(* Logix 5000 project; controller MV vendor 1 type 14 code 217 rev 31.11; software revision 31.00; part 20 of 53 *)
(* tags used below, declared in another part *)
   CheckTimeMask : INT;
   CWD : CHECKWORD_FLAGS;
   Delphi_Does_Eng_Func : BOOL;
   MC_CH1_DR2 : PlantItem;   // CH1_DR2
   MC_CH1_DT1 : PlantItem;   // CH1_DT1
   MC_CH1_DT2 : PlantItem;   // CH1_DT2
   MC_CH1_LF1 : PlantItem;   // CH1_LF1
   MC_CH1_PR1 : PlantItem;   // CH1_PR1
   MC_CH2_R1 : PlantItem;   // CH2_R1
   MC_CH2_R1R : PlantItem;   // CH2_R1R
   MC_CH2_R2 : PlantItem;   // CH2_R2
   MC_CH2_R2R : PlantItem;   // CH2_R2R
   MC_CH2_R3 : PlantItem;   // CH2_R3
   MC_CH2_R4 : PlantItem;   // CH2_R4
   MC_CH2_R5 : PlantItem;   // CH2_R5
   MC_CH2_R6 : PlantItem;   // CH2_R6
   MC_N255 : INT[255];   // CHECKWORDS Plant item checkword s
   TempChecktime : DINT;
(* MC_Common, continued *)

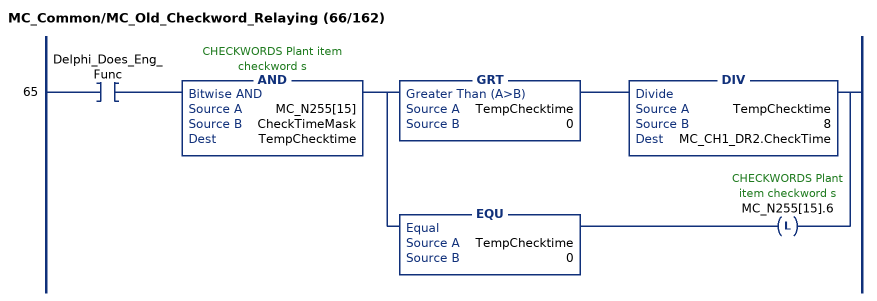
   [picture p337: MC_Common/MC_Old_Checkword_Relaying rungs 65-65]
   65: XIC(Delphi_Does_Eng_Func)AND(MC_N255[15],CheckTimeMask,TempChecktime)[GRT(TempChecktime,0) DIV(TempChecktime,8,MC_CH1_DR2.CheckTime) ,EQU(TempChecktime,0) OTL(MC_N255[15].6) ];
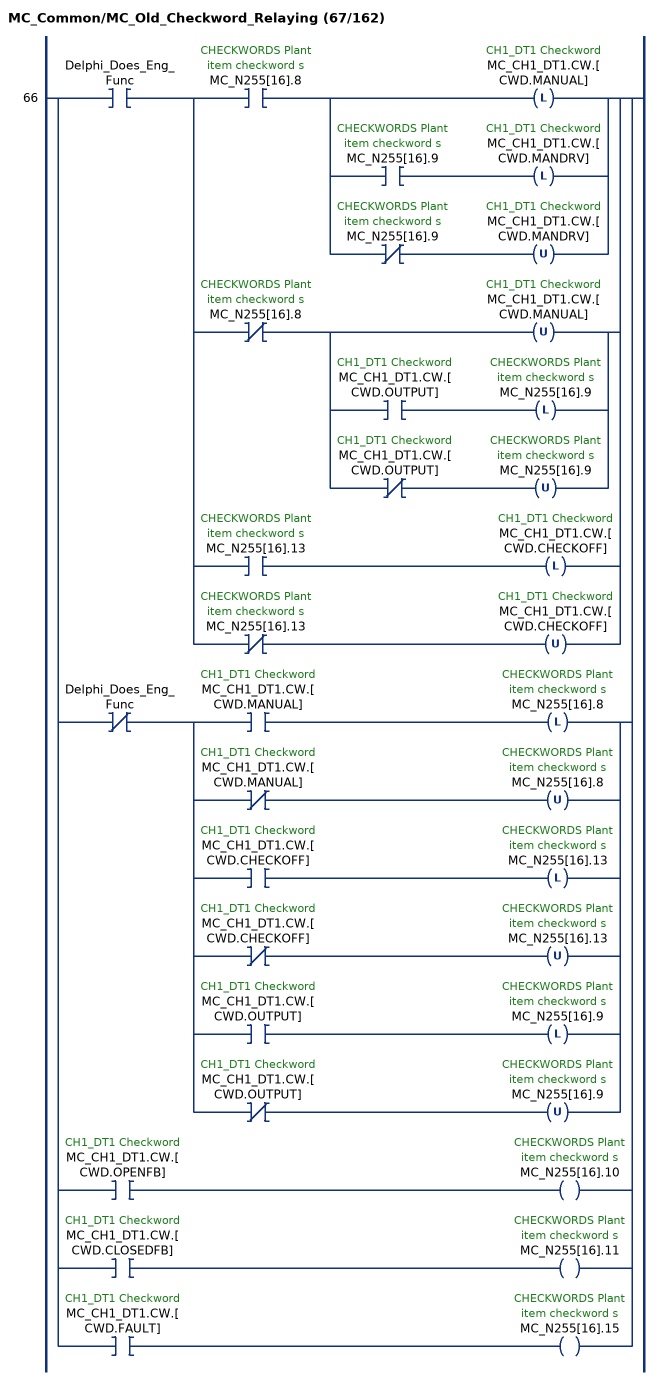
   66: [XIC(Delphi_Does_Eng_Func) [[XIC(MC_N255[16].8) [OTL(MC_CH1_DT1.CW.[CWD.MANUAL]) ,XIC(MC_N255[16].9) OTL(MC_CH1_DT1.CW.[CWD.MANDRV]) ,XIO(MC_N255[16].9) OTU(MC_CH1_DT1.CW.[CWD.MANDRV]) ] ,XIO(MC_N255[16].8) [OTU(MC_CH1_DT1.CW.[CWD.MANUAL]) ,[XIC(MC_CH1_DT1.CW.[CWD.OUTPUT]) OTL(MC_N255[16].9) ,XIO(MC_CH1_DT1.CW.[CWD.OUTPUT]) OTU(MC_N255[16].9) ] ] ] ,[XIC(MC_N255[16].13) OTL(MC_CH1_DT1.CW.[CWD.CHECKOFF]) ,XIO(MC_N255[16].13) OTU(MC_CH1_DT1.CW.[CWD.CHECKOFF]) ] ] ,XIO(Delphi_Does_Eng_Func) [[XIC(MC_CH1_DT1.CW.[CWD.MANUAL]) OTL(MC_N255[16].8) ,XIO(MC_CH1_DT1.CW.[CWD.MANUAL]) OTU(MC_N255[16].8) ] ,[XIC(MC_CH1_DT1.CW.[CWD.CHECKOFF]) OTL(MC_N255[16].13) ,XIO(MC_CH1_DT1.CW.[CWD.CHECKOFF]) OTU(MC_N255[16].13) ] ,[XIC(MC_CH1_DT1.CW.[CWD.OUTPUT]) OTL(MC_N255[16].9) ,XIO(MC_CH1_DT1.CW.[CWD.OUTPUT]) OTU(MC_N255[16].9) ] ] ,XIC(MC_CH1_DT1.CW.[CWD.OPENFB]) OTE(MC_N255[16].10) ,XIC(MC_CH1_DT1.CW.[CWD.CLOSEDFB]) OTE(MC_N255[16].11) ,XIC(MC_CH1_DT1.CW.[CWD.FAULT]) OTE(MC_N255[16].15) ];
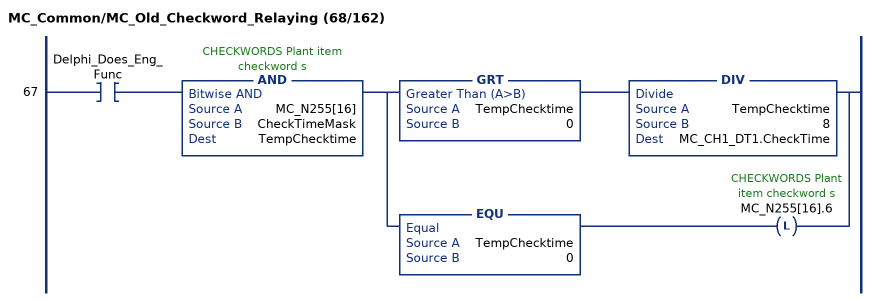
   67: XIC(Delphi_Does_Eng_Func)AND(MC_N255[16],CheckTimeMask,TempChecktime)[GRT(TempChecktime,0) DIV(TempChecktime,8,MC_CH1_DT1.CheckTime) ,EQU(TempChecktime,0) OTL(MC_N255[16].6) ];
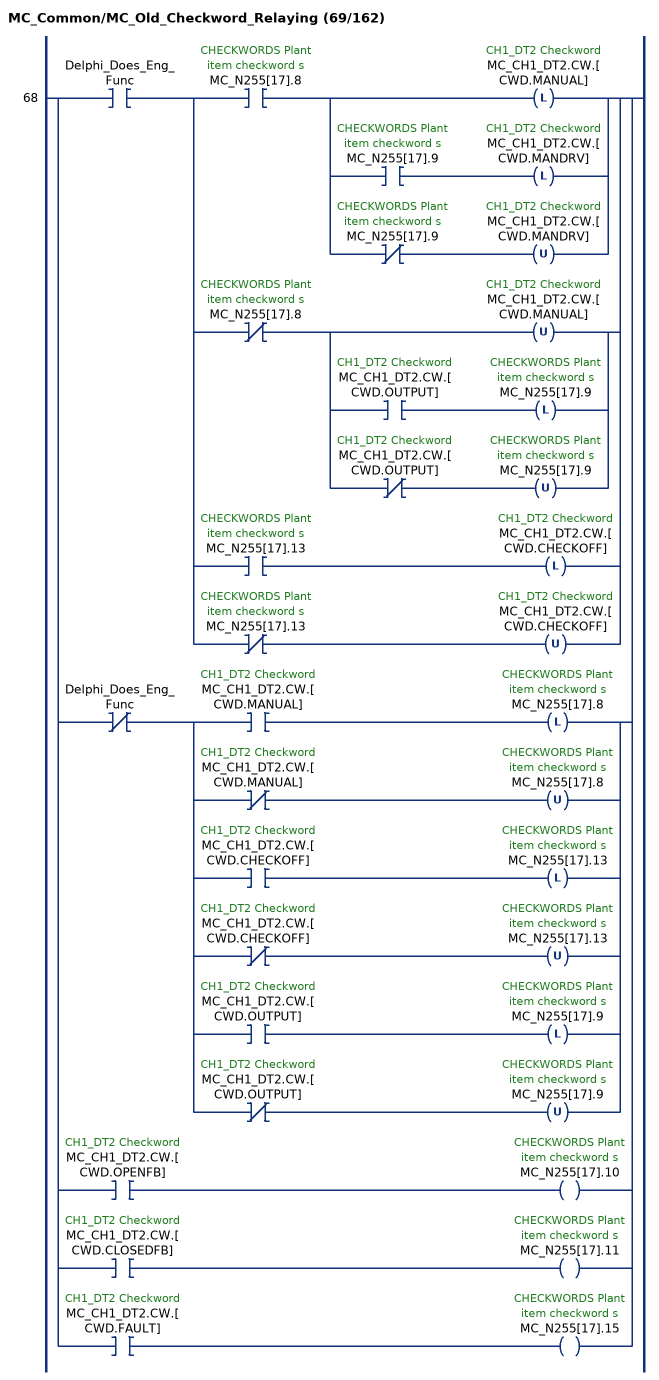
   68: [XIC(Delphi_Does_Eng_Func) [[XIC(MC_N255[17].8) [OTL(MC_CH1_DT2.CW.[CWD.MANUAL]) ,XIC(MC_N255[17].9) OTL(MC_CH1_DT2.CW.[CWD.MANDRV]) ,XIO(MC_N255[17].9) OTU(MC_CH1_DT2.CW.[CWD.MANDRV]) ] ,XIO(MC_N255[17].8) [OTU(MC_CH1_DT2.CW.[CWD.MANUAL]) ,[XIC(MC_CH1_DT2.CW.[CWD.OUTPUT]) OTL(MC_N255[17].9) ,XIO(MC_CH1_DT2.CW.[CWD.OUTPUT]) OTU(MC_N255[17].9) ] ] ] ,[XIC(MC_N255[17].13) OTL(MC_CH1_DT2.CW.[CWD.CHECKOFF]) ,XIO(MC_N255[17].13) OTU(MC_CH1_DT2.CW.[CWD.CHECKOFF]) ] ] ,XIO(Delphi_Does_Eng_Func) [[XIC(MC_CH1_DT2.CW.[CWD.MANUAL]) OTL(MC_N255[17].8) ,XIO(MC_CH1_DT2.CW.[CWD.MANUAL]) OTU(MC_N255[17].8) ] ,[XIC(MC_CH1_DT2.CW.[CWD.CHECKOFF]) OTL(MC_N255[17].13) ,XIO(MC_CH1_DT2.CW.[CWD.CHECKOFF]) OTU(MC_N255[17].13) ] ,[XIC(MC_CH1_DT2.CW.[CWD.OUTPUT]) OTL(MC_N255[17].9) ,XIO(MC_CH1_DT2.CW.[CWD.OUTPUT]) OTU(MC_N255[17].9) ] ] ,XIC(MC_CH1_DT2.CW.[CWD.OPENFB]) OTE(MC_N255[17].10) ,XIC(MC_CH1_DT2.CW.[CWD.CLOSEDFB]) OTE(MC_N255[17].11) ,XIC(MC_CH1_DT2.CW.[CWD.FAULT]) OTE(MC_N255[17].15) ];
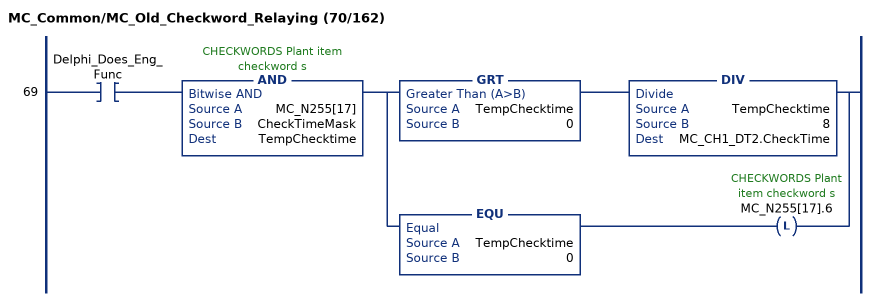
   69: XIC(Delphi_Does_Eng_Func)AND(MC_N255[17],CheckTimeMask,TempChecktime)[GRT(TempChecktime,0) DIV(TempChecktime,8,MC_CH1_DT2.CheckTime) ,EQU(TempChecktime,0) OTL(MC_N255[17].6) ];
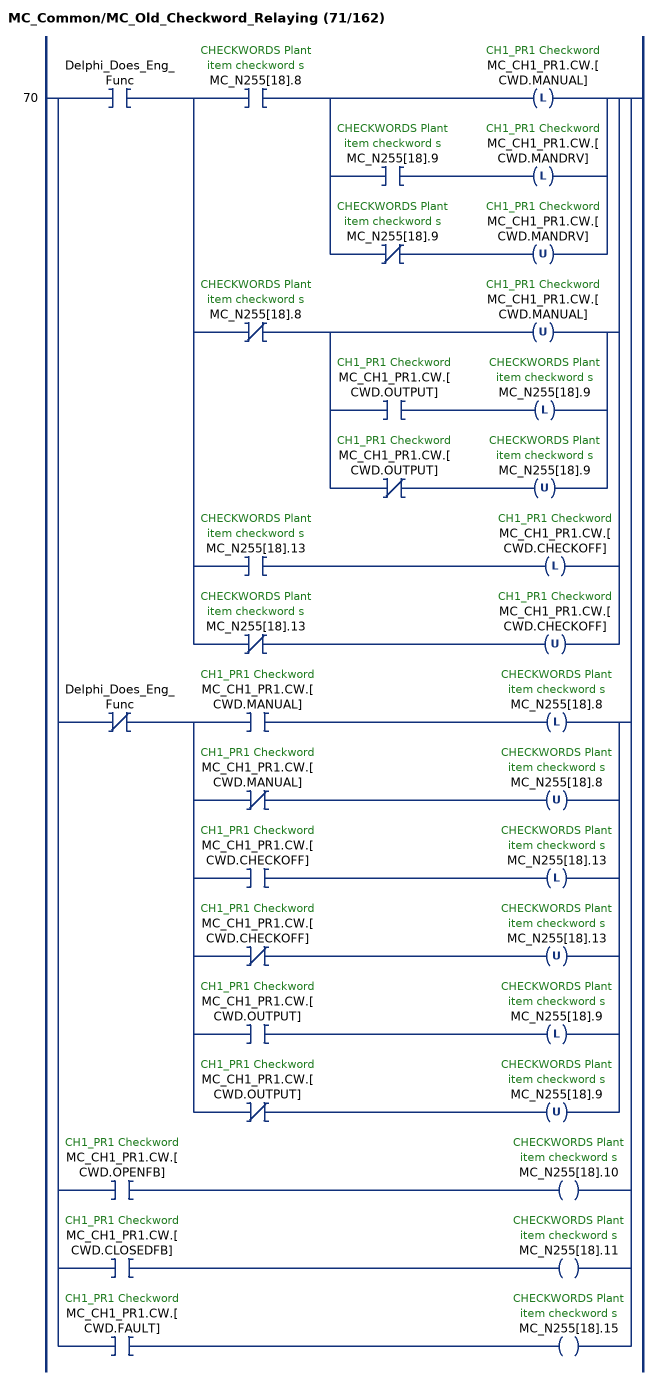
   70: [XIC(Delphi_Does_Eng_Func) [[XIC(MC_N255[18].8) [OTL(MC_CH1_PR1.CW.[CWD.MANUAL]) ,XIC(MC_N255[18].9) OTL(MC_CH1_PR1.CW.[CWD.MANDRV]) ,XIO(MC_N255[18].9) OTU(MC_CH1_PR1.CW.[CWD.MANDRV]) ] ,XIO(MC_N255[18].8) [OTU(MC_CH1_PR1.CW.[CWD.MANUAL]) ,[XIC(MC_CH1_PR1.CW.[CWD.OUTPUT]) OTL(MC_N255[18].9) ,XIO(MC_CH1_PR1.CW.[CWD.OUTPUT]) OTU(MC_N255[18].9) ] ] ] ,[XIC(MC_N255[18].13) OTL(MC_CH1_PR1.CW.[CWD.CHECKOFF]) ,XIO(MC_N255[18].13) OTU(MC_CH1_PR1.CW.[CWD.CHECKOFF]) ] ] ,XIO(Delphi_Does_Eng_Func) [[XIC(MC_CH1_PR1.CW.[CWD.MANUAL]) OTL(MC_N255[18].8) ,XIO(MC_CH1_PR1.CW.[CWD.MANUAL]) OTU(MC_N255[18].8) ] ,[XIC(MC_CH1_PR1.CW.[CWD.CHECKOFF]) OTL(MC_N255[18].13) ,XIO(MC_CH1_PR1.CW.[CWD.CHECKOFF]) OTU(MC_N255[18].13) ] ,[XIC(MC_CH1_PR1.CW.[CWD.OUTPUT]) OTL(MC_N255[18].9) ,XIO(MC_CH1_PR1.CW.[CWD.OUTPUT]) OTU(MC_N255[18].9) ] ] ,XIC(MC_CH1_PR1.CW.[CWD.OPENFB]) OTE(MC_N255[18].10) ,XIC(MC_CH1_PR1.CW.[CWD.CLOSEDFB]) OTE(MC_N255[18].11) ,XIC(MC_CH1_PR1.CW.[CWD.FAULT]) OTE(MC_N255[18].15) ];
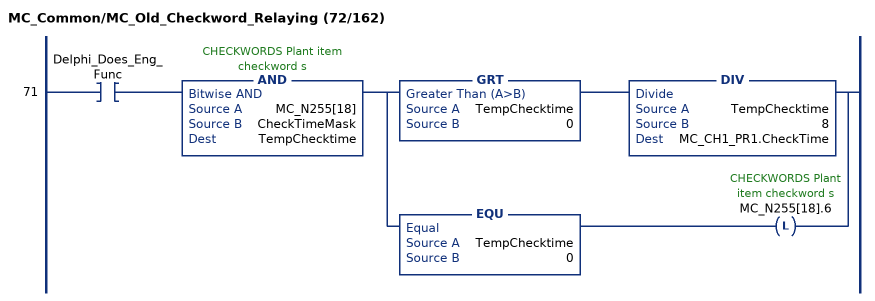
   71: XIC(Delphi_Does_Eng_Func)AND(MC_N255[18],CheckTimeMask,TempChecktime)[GRT(TempChecktime,0) DIV(TempChecktime,8,MC_CH1_PR1.CheckTime) ,EQU(TempChecktime,0) OTL(MC_N255[18].6) ];
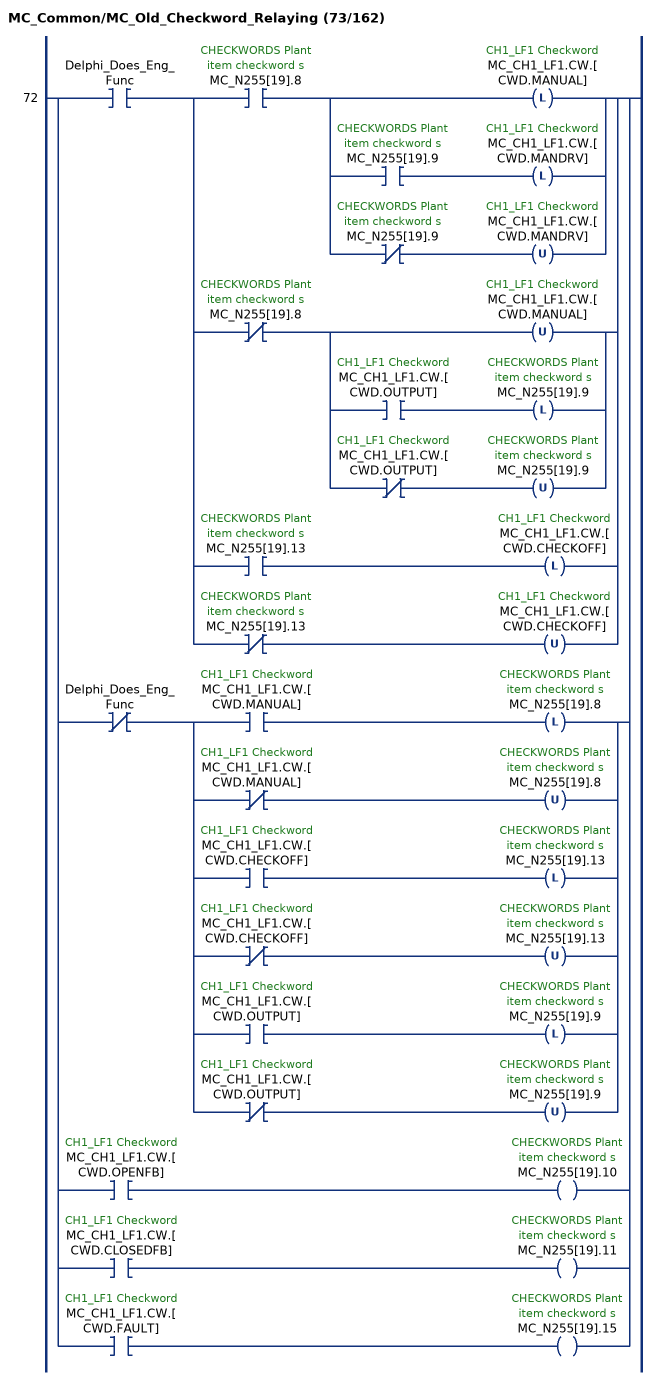
   72: [XIC(Delphi_Does_Eng_Func) [[XIC(MC_N255[19].8) [OTL(MC_CH1_LF1.CW.[CWD.MANUAL]) ,XIC(MC_N255[19].9) OTL(MC_CH1_LF1.CW.[CWD.MANDRV]) ,XIO(MC_N255[19].9) OTU(MC_CH1_LF1.CW.[CWD.MANDRV]) ] ,XIO(MC_N255[19].8) [OTU(MC_CH1_LF1.CW.[CWD.MANUAL]) ,[XIC(MC_CH1_LF1.CW.[CWD.OUTPUT]) OTL(MC_N255[19].9) ,XIO(MC_CH1_LF1.CW.[CWD.OUTPUT]) OTU(MC_N255[19].9) ] ] ] ,[XIC(MC_N255[19].13) OTL(MC_CH1_LF1.CW.[CWD.CHECKOFF]) ,XIO(MC_N255[19].13) OTU(MC_CH1_LF1.CW.[CWD.CHECKOFF]) ] ] ,XIO(Delphi_Does_Eng_Func) [[XIC(MC_CH1_LF1.CW.[CWD.MANUAL]) OTL(MC_N255[19].8) ,XIO(MC_CH1_LF1.CW.[CWD.MANUAL]) OTU(MC_N255[19].8) ] ,[XIC(MC_CH1_LF1.CW.[CWD.CHECKOFF]) OTL(MC_N255[19].13) ,XIO(MC_CH1_LF1.CW.[CWD.CHECKOFF]) OTU(MC_N255[19].13) ] ,[XIC(MC_CH1_LF1.CW.[CWD.OUTPUT]) OTL(MC_N255[19].9) ,XIO(MC_CH1_LF1.CW.[CWD.OUTPUT]) OTU(MC_N255[19].9) ] ] ,XIC(MC_CH1_LF1.CW.[CWD.OPENFB]) OTE(MC_N255[19].10) ,XIC(MC_CH1_LF1.CW.[CWD.CLOSEDFB]) OTE(MC_N255[19].11) ,XIC(MC_CH1_LF1.CW.[CWD.FAULT]) OTE(MC_N255[19].15) ];
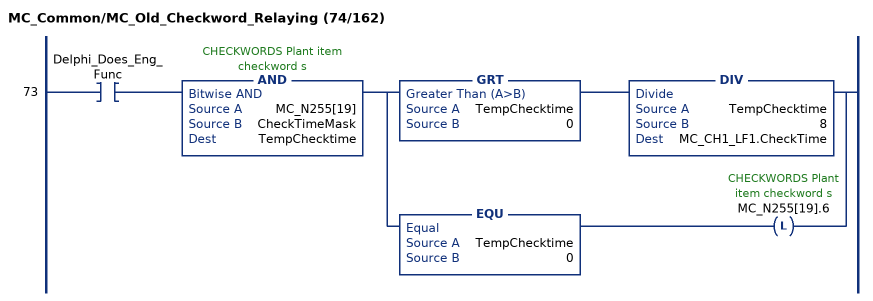
   73: XIC(Delphi_Does_Eng_Func)AND(MC_N255[19],CheckTimeMask,TempChecktime)[GRT(TempChecktime,0) DIV(TempChecktime,8,MC_CH1_LF1.CheckTime) ,EQU(TempChecktime,0) OTL(MC_N255[19].6) ];
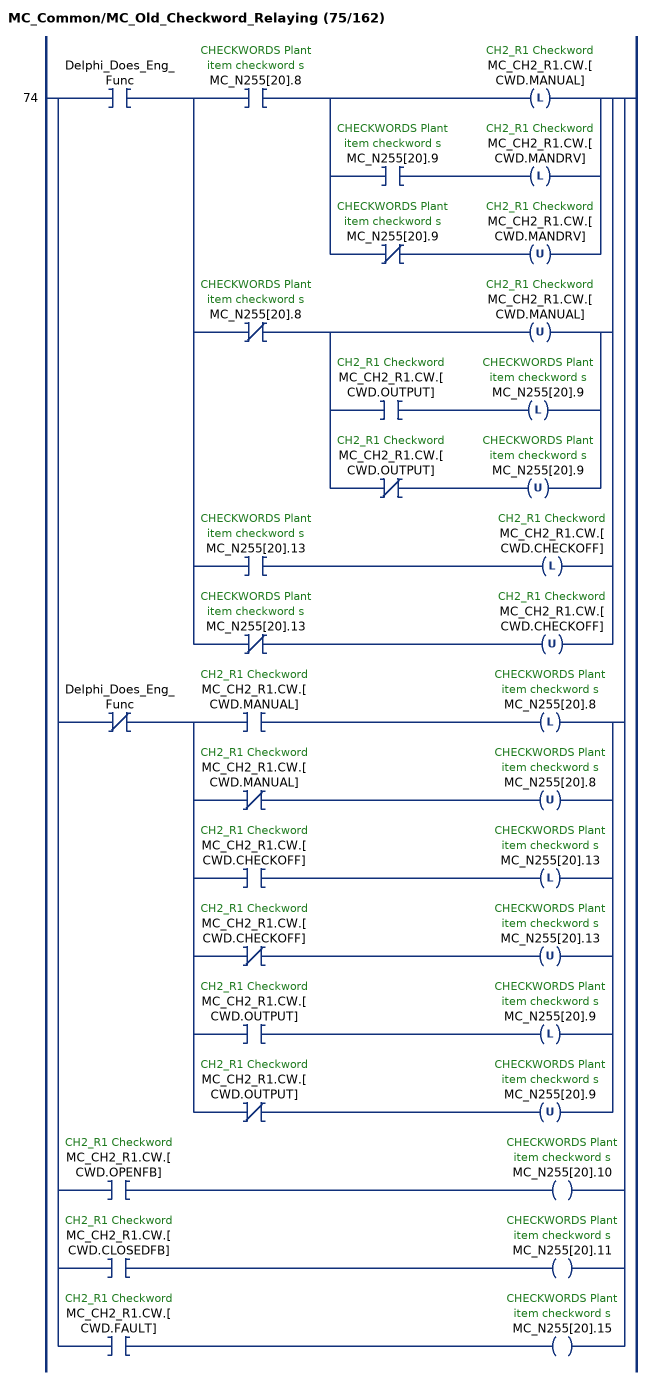
   74: [XIC(Delphi_Does_Eng_Func) [[XIC(MC_N255[20].8) [OTL(MC_CH2_R1.CW.[CWD.MANUAL]) ,XIC(MC_N255[20].9) OTL(MC_CH2_R1.CW.[CWD.MANDRV]) ,XIO(MC_N255[20].9) OTU(MC_CH2_R1.CW.[CWD.MANDRV]) ] ,XIO(MC_N255[20].8) [OTU(MC_CH2_R1.CW.[CWD.MANUAL]) ,[XIC(MC_CH2_R1.CW.[CWD.OUTPUT]) OTL(MC_N255[20].9) ,XIO(MC_CH2_R1.CW.[CWD.OUTPUT]) OTU(MC_N255[20].9) ] ] ] ,[XIC(MC_N255[20].13) OTL(MC_CH2_R1.CW.[CWD.CHECKOFF]) ,XIO(MC_N255[20].13) OTU(MC_CH2_R1.CW.[CWD.CHECKOFF]) ] ] ,XIO(Delphi_Does_Eng_Func) [[XIC(MC_CH2_R1.CW.[CWD.MANUAL]) OTL(MC_N255[20].8) ,XIO(MC_CH2_R1.CW.[CWD.MANUAL]) OTU(MC_N255[20].8) ] ,[XIC(MC_CH2_R1.CW.[CWD.CHECKOFF]) OTL(MC_N255[20].13) ,XIO(MC_CH2_R1.CW.[CWD.CHECKOFF]) OTU(MC_N255[20].13) ] ,[XIC(MC_CH2_R1.CW.[CWD.OUTPUT]) OTL(MC_N255[20].9) ,XIO(MC_CH2_R1.CW.[CWD.OUTPUT]) OTU(MC_N255[20].9) ] ] ,XIC(MC_CH2_R1.CW.[CWD.OPENFB]) OTE(MC_N255[20].10) ,XIC(MC_CH2_R1.CW.[CWD.CLOSEDFB]) OTE(MC_N255[20].11) ,XIC(MC_CH2_R1.CW.[CWD.FAULT]) OTE(MC_N255[20].15) ];
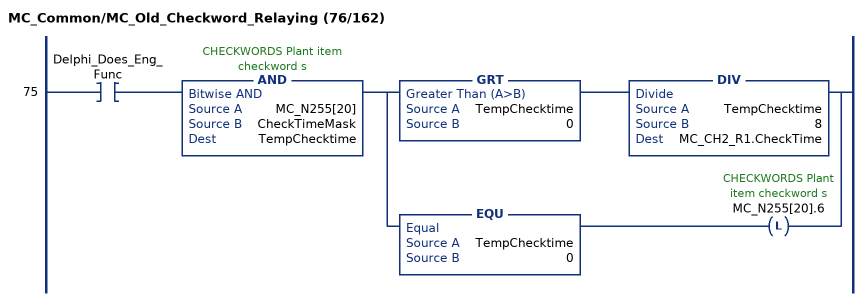
   75: XIC(Delphi_Does_Eng_Func)AND(MC_N255[20],CheckTimeMask,TempChecktime)[GRT(TempChecktime,0) DIV(TempChecktime,8,MC_CH2_R1.CheckTime) ,EQU(TempChecktime,0) OTL(MC_N255[20].6) ];
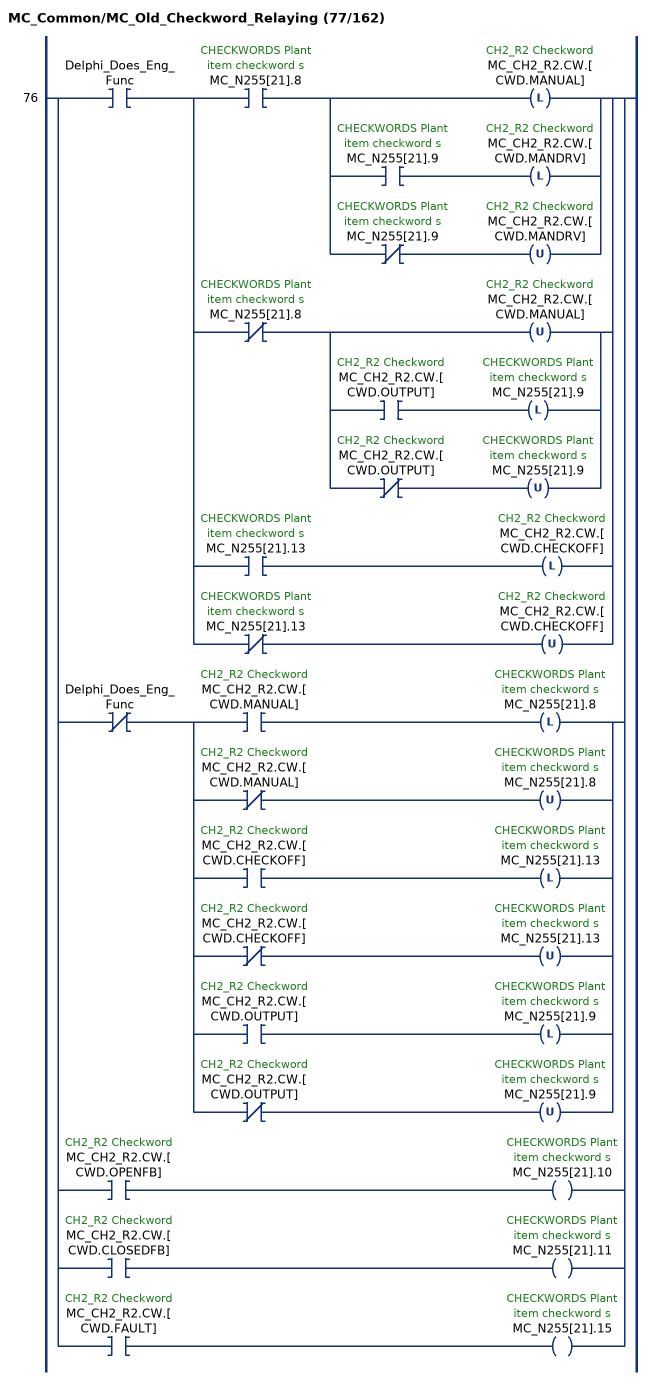
   76: [XIC(Delphi_Does_Eng_Func) [[XIC(MC_N255[21].8) [OTL(MC_CH2_R2.CW.[CWD.MANUAL]) ,XIC(MC_N255[21].9) OTL(MC_CH2_R2.CW.[CWD.MANDRV]) ,XIO(MC_N255[21].9) OTU(MC_CH2_R2.CW.[CWD.MANDRV]) ] ,XIO(MC_N255[21].8) [OTU(MC_CH2_R2.CW.[CWD.MANUAL]) ,[XIC(MC_CH2_R2.CW.[CWD.OUTPUT]) OTL(MC_N255[21].9) ,XIO(MC_CH2_R2.CW.[CWD.OUTPUT]) OTU(MC_N255[21].9) ] ] ] ,[XIC(MC_N255[21].13) OTL(MC_CH2_R2.CW.[CWD.CHECKOFF]) ,XIO(MC_N255[21].13) OTU(MC_CH2_R2.CW.[CWD.CHECKOFF]) ] ] ,XIO(Delphi_Does_Eng_Func) [[XIC(MC_CH2_R2.CW.[CWD.MANUAL]) OTL(MC_N255[21].8) ,XIO(MC_CH2_R2.CW.[CWD.MANUAL]) OTU(MC_N255[21].8) ] ,[XIC(MC_CH2_R2.CW.[CWD.CHECKOFF]) OTL(MC_N255[21].13) ,XIO(MC_CH2_R2.CW.[CWD.CHECKOFF]) OTU(MC_N255[21].13) ] ,[XIC(MC_CH2_R2.CW.[CWD.OUTPUT]) OTL(MC_N255[21].9) ,XIO(MC_CH2_R2.CW.[CWD.OUTPUT]) OTU(MC_N255[21].9) ] ] ,XIC(MC_CH2_R2.CW.[CWD.OPENFB]) OTE(MC_N255[21].10) ,XIC(MC_CH2_R2.CW.[CWD.CLOSEDFB]) OTE(MC_N255[21].11) ,XIC(MC_CH2_R2.CW.[CWD.FAULT]) OTE(MC_N255[21].15) ];
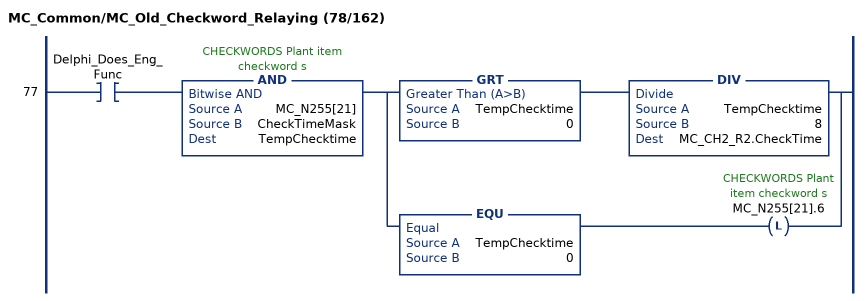
   77: XIC(Delphi_Does_Eng_Func)AND(MC_N255[21],CheckTimeMask,TempChecktime)[GRT(TempChecktime,0) DIV(TempChecktime,8,MC_CH2_R2.CheckTime) ,EQU(TempChecktime,0) OTL(MC_N255[21].6) ];
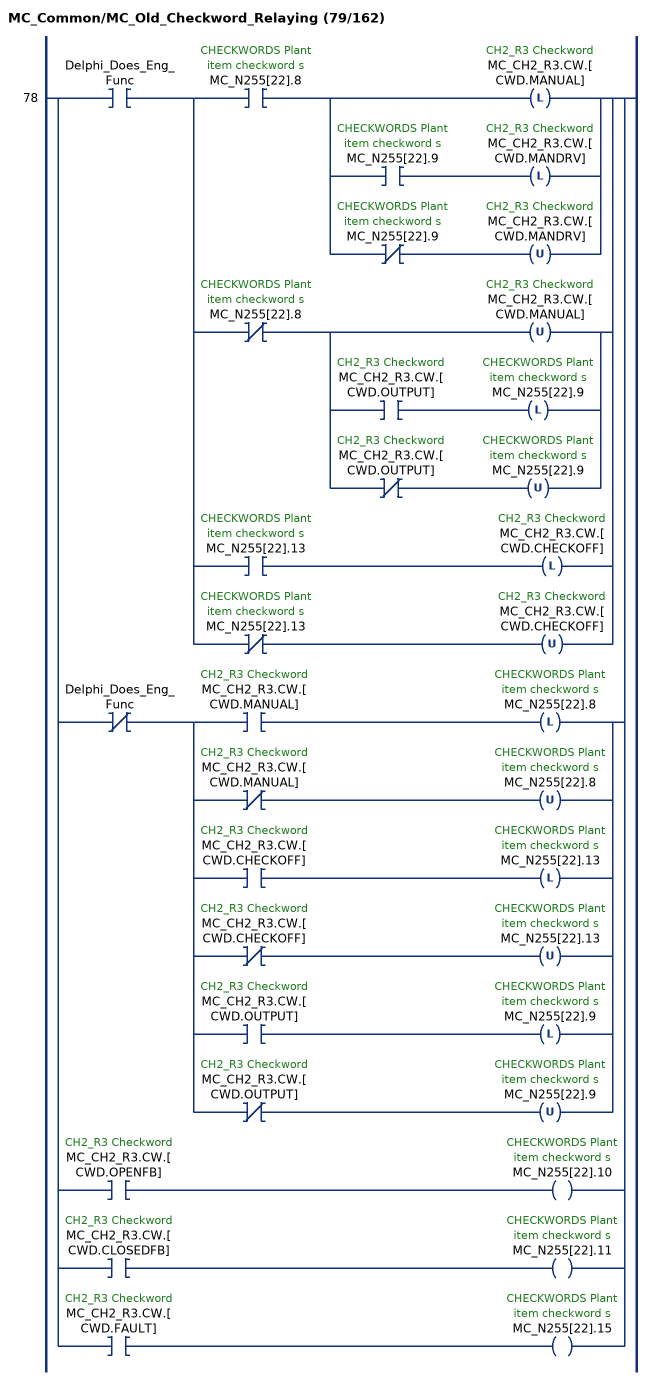
   78: [XIC(Delphi_Does_Eng_Func) [[XIC(MC_N255[22].8) [OTL(MC_CH2_R3.CW.[CWD.MANUAL]) ,XIC(MC_N255[22].9) OTL(MC_CH2_R3.CW.[CWD.MANDRV]) ,XIO(MC_N255[22].9) OTU(MC_CH2_R3.CW.[CWD.MANDRV]) ] ,XIO(MC_N255[22].8) [OTU(MC_CH2_R3.CW.[CWD.MANUAL]) ,[XIC(MC_CH2_R3.CW.[CWD.OUTPUT]) OTL(MC_N255[22].9) ,XIO(MC_CH2_R3.CW.[CWD.OUTPUT]) OTU(MC_N255[22].9) ] ] ] ,[XIC(MC_N255[22].13) OTL(MC_CH2_R3.CW.[CWD.CHECKOFF]) ,XIO(MC_N255[22].13) OTU(MC_CH2_R3.CW.[CWD.CHECKOFF]) ] ] ,XIO(Delphi_Does_Eng_Func) [[XIC(MC_CH2_R3.CW.[CWD.MANUAL]) OTL(MC_N255[22].8) ,XIO(MC_CH2_R3.CW.[CWD.MANUAL]) OTU(MC_N255[22].8) ] ,[XIC(MC_CH2_R3.CW.[CWD.CHECKOFF]) OTL(MC_N255[22].13) ,XIO(MC_CH2_R3.CW.[CWD.CHECKOFF]) OTU(MC_N255[22].13) ] ,[XIC(MC_CH2_R3.CW.[CWD.OUTPUT]) OTL(MC_N255[22].9) ,XIO(MC_CH2_R3.CW.[CWD.OUTPUT]) OTU(MC_N255[22].9) ] ] ,XIC(MC_CH2_R3.CW.[CWD.OPENFB]) OTE(MC_N255[22].10) ,XIC(MC_CH2_R3.CW.[CWD.CLOSEDFB]) OTE(MC_N255[22].11) ,XIC(MC_CH2_R3.CW.[CWD.FAULT]) OTE(MC_N255[22].15) ];
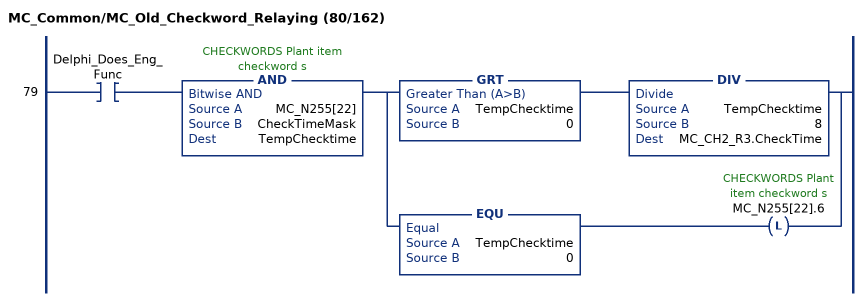
   79: XIC(Delphi_Does_Eng_Func)AND(MC_N255[22],CheckTimeMask,TempChecktime)[GRT(TempChecktime,0) DIV(TempChecktime,8,MC_CH2_R3.CheckTime) ,EQU(TempChecktime,0) OTL(MC_N255[22].6) ];
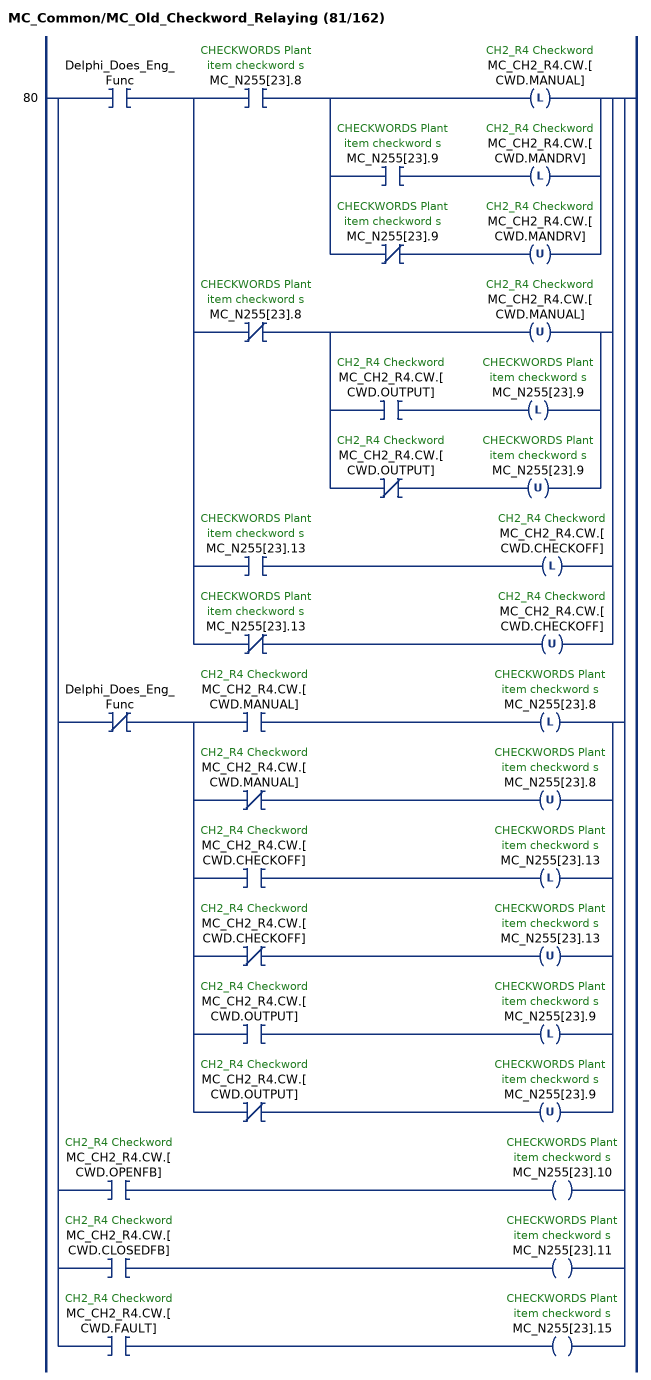
   80: [XIC(Delphi_Does_Eng_Func) [[XIC(MC_N255[23].8) [OTL(MC_CH2_R4.CW.[CWD.MANUAL]) ,XIC(MC_N255[23].9) OTL(MC_CH2_R4.CW.[CWD.MANDRV]) ,XIO(MC_N255[23].9) OTU(MC_CH2_R4.CW.[CWD.MANDRV]) ] ,XIO(MC_N255[23].8) [OTU(MC_CH2_R4.CW.[CWD.MANUAL]) ,[XIC(MC_CH2_R4.CW.[CWD.OUTPUT]) OTL(MC_N255[23].9) ,XIO(MC_CH2_R4.CW.[CWD.OUTPUT]) OTU(MC_N255[23].9) ] ] ] ,[XIC(MC_N255[23].13) OTL(MC_CH2_R4.CW.[CWD.CHECKOFF]) ,XIO(MC_N255[23].13) OTU(MC_CH2_R4.CW.[CWD.CHECKOFF]) ] ] ,XIO(Delphi_Does_Eng_Func) [[XIC(MC_CH2_R4.CW.[CWD.MANUAL]) OTL(MC_N255[23].8) ,XIO(MC_CH2_R4.CW.[CWD.MANUAL]) OTU(MC_N255[23].8) ] ,[XIC(MC_CH2_R4.CW.[CWD.CHECKOFF]) OTL(MC_N255[23].13) ,XIO(MC_CH2_R4.CW.[CWD.CHECKOFF]) OTU(MC_N255[23].13) ] ,[XIC(MC_CH2_R4.CW.[CWD.OUTPUT]) OTL(MC_N255[23].9) ,XIO(MC_CH2_R4.CW.[CWD.OUTPUT]) OTU(MC_N255[23].9) ] ] ,XIC(MC_CH2_R4.CW.[CWD.OPENFB]) OTE(MC_N255[23].10) ,XIC(MC_CH2_R4.CW.[CWD.CLOSEDFB]) OTE(MC_N255[23].11) ,XIC(MC_CH2_R4.CW.[CWD.FAULT]) OTE(MC_N255[23].15) ];
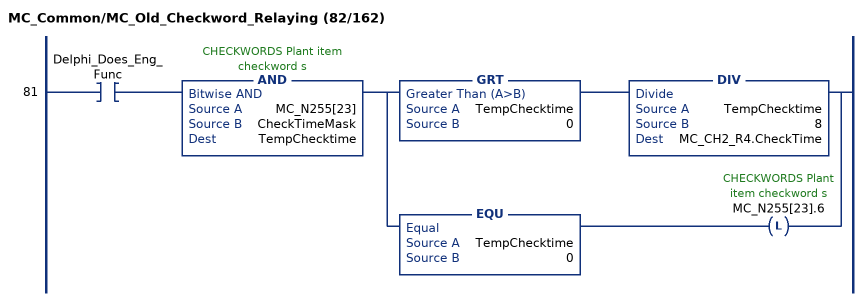
   81: XIC(Delphi_Does_Eng_Func)AND(MC_N255[23],CheckTimeMask,TempChecktime)[GRT(TempChecktime,0) DIV(TempChecktime,8,MC_CH2_R4.CheckTime) ,EQU(TempChecktime,0) OTL(MC_N255[23].6) ];
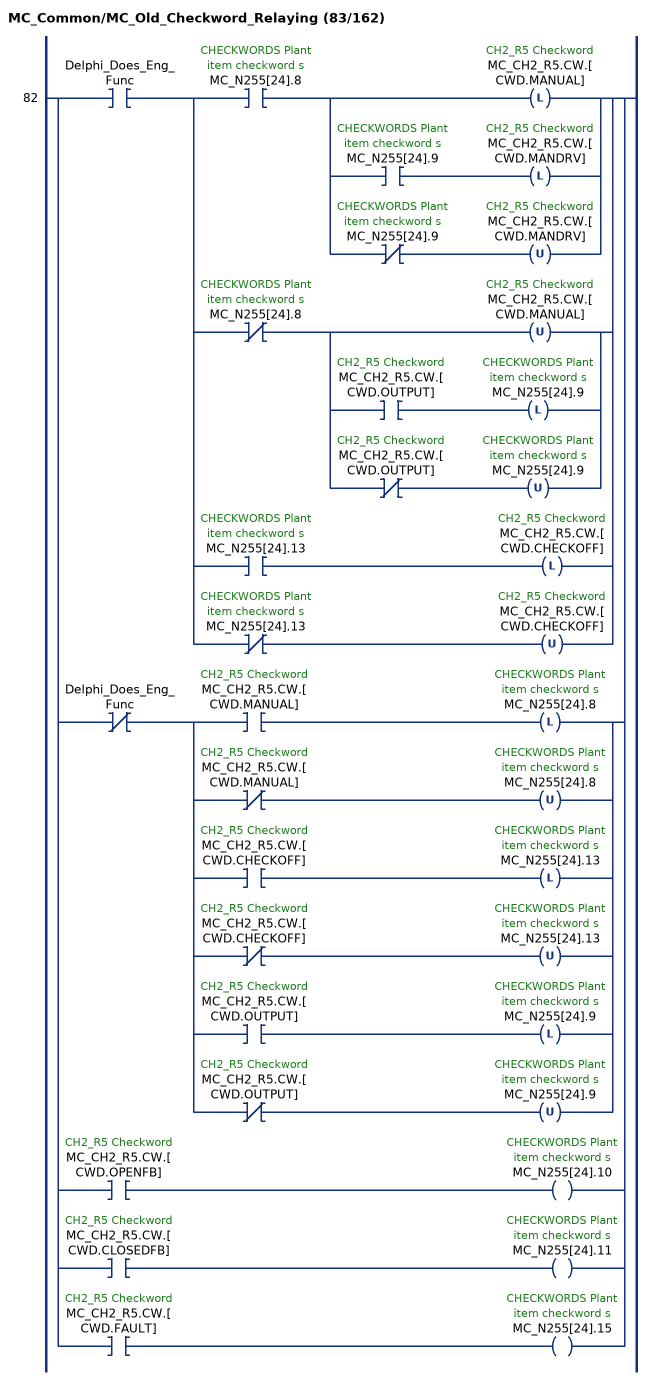
   82: [XIC(Delphi_Does_Eng_Func) [[XIC(MC_N255[24].8) [OTL(MC_CH2_R5.CW.[CWD.MANUAL]) ,XIC(MC_N255[24].9) OTL(MC_CH2_R5.CW.[CWD.MANDRV]) ,XIO(MC_N255[24].9) OTU(MC_CH2_R5.CW.[CWD.MANDRV]) ] ,XIO(MC_N255[24].8) [OTU(MC_CH2_R5.CW.[CWD.MANUAL]) ,[XIC(MC_CH2_R5.CW.[CWD.OUTPUT]) OTL(MC_N255[24].9) ,XIO(MC_CH2_R5.CW.[CWD.OUTPUT]) OTU(MC_N255[24].9) ] ] ] ,[XIC(MC_N255[24].13) OTL(MC_CH2_R5.CW.[CWD.CHECKOFF]) ,XIO(MC_N255[24].13) OTU(MC_CH2_R5.CW.[CWD.CHECKOFF]) ] ] ,XIO(Delphi_Does_Eng_Func) [[XIC(MC_CH2_R5.CW.[CWD.MANUAL]) OTL(MC_N255[24].8) ,XIO(MC_CH2_R5.CW.[CWD.MANUAL]) OTU(MC_N255[24].8) ] ,[XIC(MC_CH2_R5.CW.[CWD.CHECKOFF]) OTL(MC_N255[24].13) ,XIO(MC_CH2_R5.CW.[CWD.CHECKOFF]) OTU(MC_N255[24].13) ] ,[XIC(MC_CH2_R5.CW.[CWD.OUTPUT]) OTL(MC_N255[24].9) ,XIO(MC_CH2_R5.CW.[CWD.OUTPUT]) OTU(MC_N255[24].9) ] ] ,XIC(MC_CH2_R5.CW.[CWD.OPENFB]) OTE(MC_N255[24].10) ,XIC(MC_CH2_R5.CW.[CWD.CLOSEDFB]) OTE(MC_N255[24].11) ,XIC(MC_CH2_R5.CW.[CWD.FAULT]) OTE(MC_N255[24].15) ];
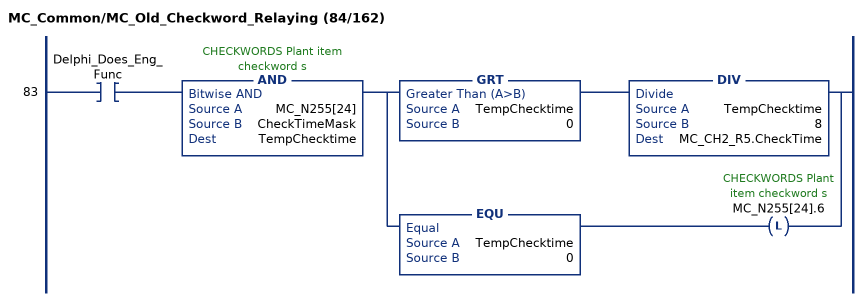
   83: XIC(Delphi_Does_Eng_Func)AND(MC_N255[24],CheckTimeMask,TempChecktime)[GRT(TempChecktime,0) DIV(TempChecktime,8,MC_CH2_R5.CheckTime) ,EQU(TempChecktime,0) OTL(MC_N255[24].6) ];
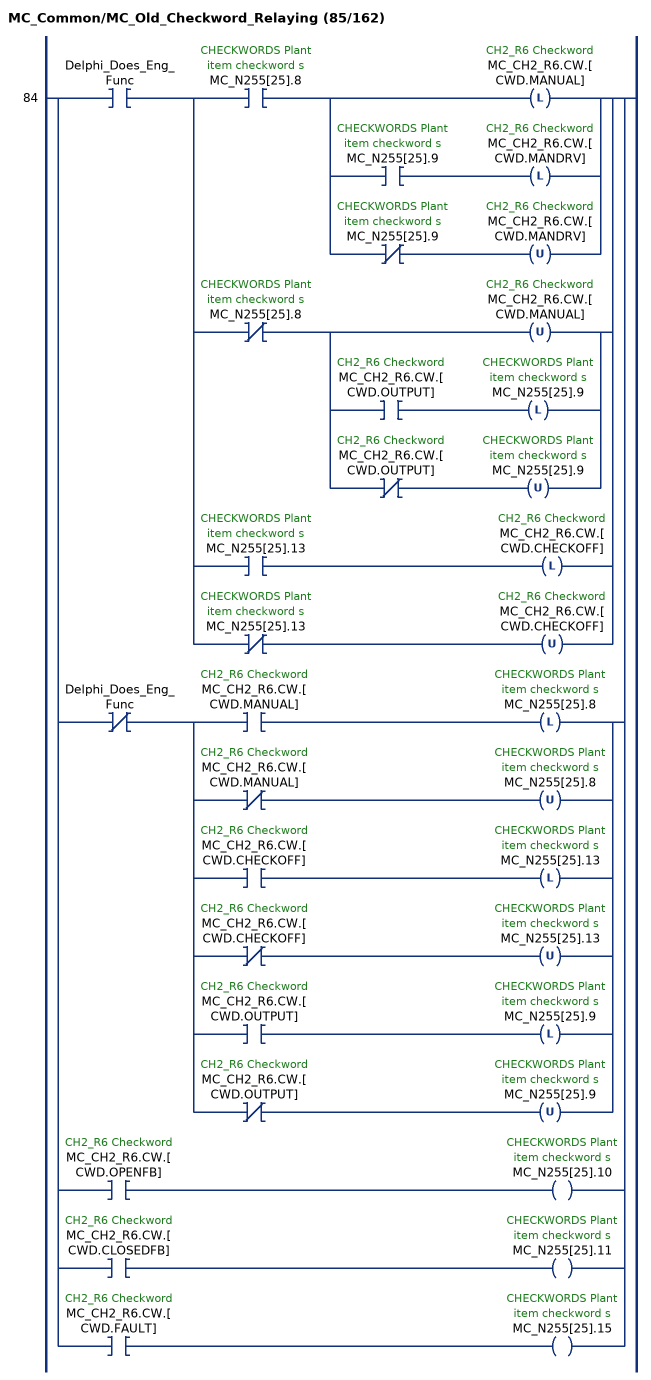
   84: [XIC(Delphi_Does_Eng_Func) [[XIC(MC_N255[25].8) [OTL(MC_CH2_R6.CW.[CWD.MANUAL]) ,XIC(MC_N255[25].9) OTL(MC_CH2_R6.CW.[CWD.MANDRV]) ,XIO(MC_N255[25].9) OTU(MC_CH2_R6.CW.[CWD.MANDRV]) ] ,XIO(MC_N255[25].8) [OTU(MC_CH2_R6.CW.[CWD.MANUAL]) ,[XIC(MC_CH2_R6.CW.[CWD.OUTPUT]) OTL(MC_N255[25].9) ,XIO(MC_CH2_R6.CW.[CWD.OUTPUT]) OTU(MC_N255[25].9) ] ] ] ,[XIC(MC_N255[25].13) OTL(MC_CH2_R6.CW.[CWD.CHECKOFF]) ,XIO(MC_N255[25].13) OTU(MC_CH2_R6.CW.[CWD.CHECKOFF]) ] ] ,XIO(Delphi_Does_Eng_Func) [[XIC(MC_CH2_R6.CW.[CWD.MANUAL]) OTL(MC_N255[25].8) ,XIO(MC_CH2_R6.CW.[CWD.MANUAL]) OTU(MC_N255[25].8) ] ,[XIC(MC_CH2_R6.CW.[CWD.CHECKOFF]) OTL(MC_N255[25].13) ,XIO(MC_CH2_R6.CW.[CWD.CHECKOFF]) OTU(MC_N255[25].13) ] ,[XIC(MC_CH2_R6.CW.[CWD.OUTPUT]) OTL(MC_N255[25].9) ,XIO(MC_CH2_R6.CW.[CWD.OUTPUT]) OTU(MC_N255[25].9) ] ] ,XIC(MC_CH2_R6.CW.[CWD.OPENFB]) OTE(MC_N255[25].10) ,XIC(MC_CH2_R6.CW.[CWD.CLOSEDFB]) OTE(MC_N255[25].11) ,XIC(MC_CH2_R6.CW.[CWD.FAULT]) OTE(MC_N255[25].15) ];
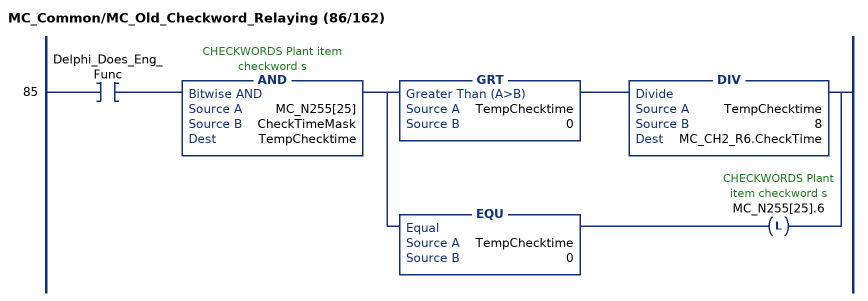
   85: XIC(Delphi_Does_Eng_Func)AND(MC_N255[25],CheckTimeMask,TempChecktime)[GRT(TempChecktime,0) DIV(TempChecktime,8,MC_CH2_R6.CheckTime) ,EQU(TempChecktime,0) OTL(MC_N255[25].6) ];
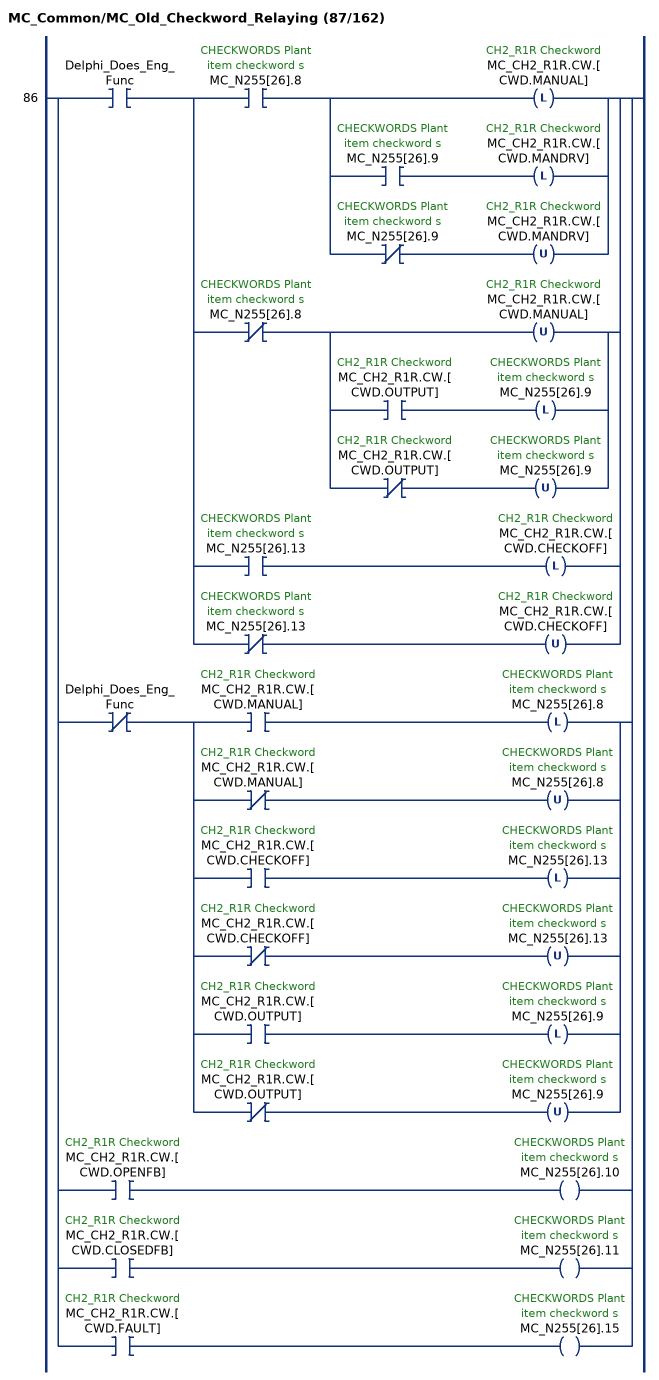
   86: [XIC(Delphi_Does_Eng_Func) [[XIC(MC_N255[26].8) [OTL(MC_CH2_R1R.CW.[CWD.MANUAL]) ,XIC(MC_N255[26].9) OTL(MC_CH2_R1R.CW.[CWD.MANDRV]) ,XIO(MC_N255[26].9) OTU(MC_CH2_R1R.CW.[CWD.MANDRV]) ] ,XIO(MC_N255[26].8) [OTU(MC_CH2_R1R.CW.[CWD.MANUAL]) ,[XIC(MC_CH2_R1R.CW.[CWD.OUTPUT]) OTL(MC_N255[26].9) ,XIO(MC_CH2_R1R.CW.[CWD.OUTPUT]) OTU(MC_N255[26].9) ] ] ] ,[XIC(MC_N255[26].13) OTL(MC_CH2_R1R.CW.[CWD.CHECKOFF]) ,XIO(MC_N255[26].13) OTU(MC_CH2_R1R.CW.[CWD.CHECKOFF]) ] ] ,XIO(Delphi_Does_Eng_Func) [[XIC(MC_CH2_R1R.CW.[CWD.MANUAL]) OTL(MC_N255[26].8) ,XIO(MC_CH2_R1R.CW.[CWD.MANUAL]) OTU(MC_N255[26].8) ] ,[XIC(MC_CH2_R1R.CW.[CWD.CHECKOFF]) OTL(MC_N255[26].13) ,XIO(MC_CH2_R1R.CW.[CWD.CHECKOFF]) OTU(MC_N255[26].13) ] ,[XIC(MC_CH2_R1R.CW.[CWD.OUTPUT]) OTL(MC_N255[26].9) ,XIO(MC_CH2_R1R.CW.[CWD.OUTPUT]) OTU(MC_N255[26].9) ] ] ,XIC(MC_CH2_R1R.CW.[CWD.OPENFB]) OTE(MC_N255[26].10) ,XIC(MC_CH2_R1R.CW.[CWD.CLOSEDFB]) OTE(MC_N255[26].11) ,XIC(MC_CH2_R1R.CW.[CWD.FAULT]) OTE(MC_N255[26].15) ];
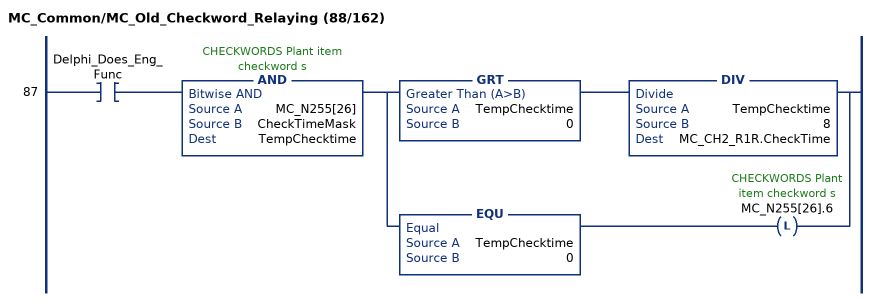
   87: XIC(Delphi_Does_Eng_Func)AND(MC_N255[26],CheckTimeMask,TempChecktime)[GRT(TempChecktime,0) DIV(TempChecktime,8,MC_CH2_R1R.CheckTime) ,EQU(TempChecktime,0) OTL(MC_N255[26].6) ];
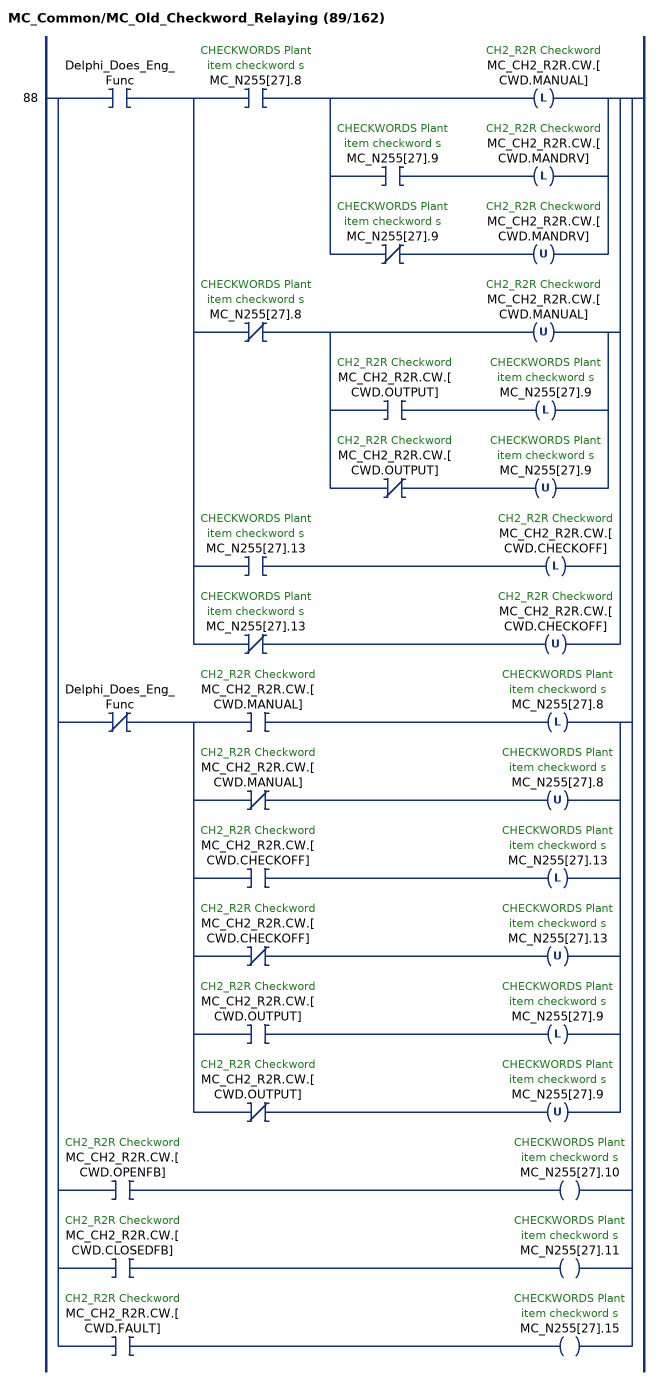
   88: [XIC(Delphi_Does_Eng_Func) [[XIC(MC_N255[27].8) [OTL(MC_CH2_R2R.CW.[CWD.MANUAL]) ,XIC(MC_N255[27].9) OTL(MC_CH2_R2R.CW.[CWD.MANDRV]) ,XIO(MC_N255[27].9) OTU(MC_CH2_R2R.CW.[CWD.MANDRV]) ] ,XIO(MC_N255[27].8) [OTU(MC_CH2_R2R.CW.[CWD.MANUAL]) ,[XIC(MC_CH2_R2R.CW.[CWD.OUTPUT]) OTL(MC_N255[27].9) ,XIO(MC_CH2_R2R.CW.[CWD.OUTPUT]) OTU(MC_N255[27].9) ] ] ] ,[XIC(MC_N255[27].13) OTL(MC_CH2_R2R.CW.[CWD.CHECKOFF]) ,XIO(MC_N255[27].13) OTU(MC_CH2_R2R.CW.[CWD.CHECKOFF]) ] ] ,XIO(Delphi_Does_Eng_Func) [[XIC(MC_CH2_R2R.CW.[CWD.MANUAL]) OTL(MC_N255[27].8) ,XIO(MC_CH2_R2R.CW.[CWD.MANUAL]) OTU(MC_N255[27].8) ] ,[XIC(MC_CH2_R2R.CW.[CWD.CHECKOFF]) OTL(MC_N255[27].13) ,XIO(MC_CH2_R2R.CW.[CWD.CHECKOFF]) OTU(MC_N255[27].13) ] ,[XIC(MC_CH2_R2R.CW.[CWD.OUTPUT]) OTL(MC_N255[27].9) ,XIO(MC_CH2_R2R.CW.[CWD.OUTPUT]) OTU(MC_N255[27].9) ] ] ,XIC(MC_CH2_R2R.CW.[CWD.OPENFB]) OTE(MC_N255[27].10) ,XIC(MC_CH2_R2R.CW.[CWD.CLOSEDFB]) OTE(MC_N255[27].11) ,XIC(MC_CH2_R2R.CW.[CWD.FAULT]) OTE(MC_N255[27].15) ];
